VERSION : 0.1
   VAR_INPUT
      Nr_Ost_Elementu : Int;   // Numer ostatniego elementu, dla ktorego wykonywana jest klasa
      Nr_Plc : Byte;
   END_VAR
   VAR_TEMP
      i : Int;
   END_VAR
BEGIN
   FOR #i := 1 TO #Nr_Ost_Elementu BY 1 DO
       REGION Opisy bitow sygnalow: bRoz,bSym,bSt,bSt_1,bTrP
           //bRoz - ROZKAZ OPERATORA - DB322.DBW10 - WORD
           //bRozB1
           //"DB322_DV1".DV1[#i].bRoZB1.%X0 - Tryb pracy: 0-Zdalny reczny; 1-Zdalny auto
           //"DB322_DV1".DV1[#i].bRoZB1.%X1 - Symulacja wejsc urz: 0-Wylaczona; 1-Zalaczona
           //"DB322_DV1".DV1[#i].bRoZB1.%X2 - Praca z wyjsciami urz: 0-Wylaczona; 1-Zalaczona
           //"DB322_DV1".DV1[#i].bRoZB1.%X3 - Sterowanie urz. w tr. Zdalnym-Man: 0-Wylacz; 1-Zalacz
           //"DB322_DV1".DV1[#i].bRoZB1.%X4 - Sterowanie kier. w tr. Zdalnym-Man: 0-Lewa; 1-Prawo
           //"DB322_DV1".DV1[#i].bRoZB1.%X5 - Rezerwa
           //"DB322_DV1".DV1[#i].bRoZB1.%X6 - Monitoring potwierdzen zal/wyl: 0-Wylaczone; 1-Zalaczone
           //"DB322_DV1".DV1[#i].bRoZB1.%X7 - Rezerwa
           //bRozB2
           //"DB322_DV1".DV1[#i].bRoZB2.%X0 - Kasuj awarie (impuls)
           //"DB322_DV1".DV1[#i].bRoZB2.%X1-X7 - Rezerwa (impuls)
           //
           //bSym - SYM WEJSCIA - DB322.DBW12 - WORD
           //"DB322_DV1".DV1[#i].bSym.%X0 - Aktywacja urz. w systemie (ustawiany tylko z programu)
           //"DB322_DV1".DV1[#i].bSym.%X1 - Sterowanie urz. w tr. Zdalnym-Auto: 0-Wylacz; 1-Zalacz
           //"DB322_DV1".DV1[#i].bSym.%X2 - Potwierdzenie zalaczenia/otwarcia
           //"DB322_DV1".DV1[#i].bSym.%X3 - Potwierdzenie wylaczenia/zamkniecia
           //"DB322_DV1".DV1[#i].bSym.%X4 - Potwierdzenie gotowosci
           //"DB322_DV1".DV1[#i].bSym.%X5 - Tryb sterowania: 0-Zdalne z PC; 1-Lokalne z elewacji szafy
           //"DB322_DV1".DV1[#i].bSym.%X6 - Tryb remontowy (z wylacznika): 0-Brak; 1-Aktywny
           //"DB322_DV1".DV1[#i].bSym.%X7 - Awaria zewnetrzna: 0-Brak; 1-Aktywny
           //"DB322_DV1".DV1[#i].bSym.%X8 - Blokada zmiany tr. zdalnego z Auto na Man: 0-Brak; 1-Aktywna
           //"DB322_DV1".DV1[#i].bSym.%X9 - Interlock w trybie Zdalnym-Auto: 0-Brak; 1-Aktywny
           //"DB322_DV1".DV1[#i].bSym.%X10-X15 - Rezerwa
           //
           //bSt_Tryb - STAN - DB322.DBW14 - WORD
           //"DB322_DV1".DV1[#i].bSt_Tryb.%X0 - Awaria od braku potwierdzen: 0-Nieaktywna; 1-Aktywna
           //"DB322_DV1".DV1[#i].bSt_Tryb.%X1 - Awaria od braku gotowosci: 0-Nieaktywna; 1-Aktywna
           //"DB322_DV1".DV1[#i].bSt_Tryb.%X2 - Awaria zewnetzrna: 0-Nieaktywna; 1-Aktywna
           //"DB322_DV1".DV1[#i].bSt_Tryb.%X3-X6 - Awaria rezerwa
           //"DB322_DV1".DV1[#i].bSt_Tryb.%X7 - Monitoring potwierdzen: 0-Wylaczony; 1-Zalaczony
           //"DB322_DV1".DV1[#i].bSt_Tryb.%X8 - Urzadzenie aktywowane
           //"DB322_DV1".DV1[#i].bSt_Tryb.%X9 - Blokada zmaiany tr. zdalnego z Auto na Man: 0-Brak; 1-Aktywna
           //"DB322_DV1".DV1[#i].bSt_Tryb.%X10 - Stan wyjścia sterującego obiekt: 0-Zamknij; 1-Otwórz
           //"DB322_DV1".DV1[#i].bSt_Tryb.%X11 - Interlock w trybie Zdalnym-Auto: 0-Brak; 1-Aktywny
           //"DB322_DV1".DV1[#i].bSt_Tryb.%X12 - Symulacja wejsc urzadzenia: 0-Wylaczona; 1-Zalaczona
           //"DB322_DV1".DV1[#i].bSt_Tryb.%X13 - Praca z wyjsciami urzadzenia: 0-Wylaczona; 1-Zalaczona
           //"DB322_DV1".DV1[#i].bSt_Tryb.%X14 - Stan urzadzenia: 0-Brak odliczania czasu do otwarcia 1-Odliczanie
           //"DB322_DV1".DV1[#i].bSt_Tryb.%X15 - Stan urzadzenia: 0-Brak odliczania czasu do zamkniecia 1-Odliczanie
           //
           //bSt_Urz - STAN - DB322.DBW16 - INT
           //"DB322_DV1".DV1[#i].bSt_Urz.%X0 - STAN(1)- Awaria zbiorcza 1-Aktywna; 0-Brak aktywnosci obiektu
           //"DB322_DV1".DV1[#i].bSt_Urz.%X1 - STAN(2)- Urzadzenie: 1-Zamkniete; 0-Inny stan
           //"DB322_DV1".DV1[#i].bSt_Urz.%X2 - STAN(4)- Urzadzenie: 1-Otwieranie; 0-Inny stan
           //"DB322_DV1".DV1[#i].bSt_Urz.%X3 - STAN(8)- Urzadzenie: 1-Otwarte; 0-Inny stan
           //"DB322_DV1".DV1[#i].bSt_Urz.%X4 - STAN(16)- Urzadzenie: 1-Zamykanie; 0-Inny stan
           //"DB322_DV1".DV1[#i].bSt_Urz.%X5 - STAN(32)- Urzadzenie: 1-Odliczanie czasu zwloki awarii; 0-Inny stan
           //"DB322_DV1".DV1[#i].bSt_Urz.%X6-X7 - STAN- Stan rezerwa
           //
           //bTrP - TRYB PRACY - DB322.DBW17 - INT
           //"DB322_DV1".DV1[#i].bTrP.%X0 - TRYB PRACY(1) - Tryb Remontowy(1): 1-Aktywny; 0-Brak aktywnosci obiektu
           //"DB322_DV1".DV1[#i].bTrP.%X1 - Tryb PRACY(2) - Tryb Sterowania: 1-Lokalny - z szafy; 0-Inny stan
           //"DB322_DV1".DV1[#i].bTrP.%X2 - TRYB PRACY(4) - Tryb Sterowania Zdalnego: 1-Zdalny Reczny; 0-Inny stan
           //"DB322_DV1".DV1[#i].bTrP.%X3 - TRYB PRACY(8) - Tryb Sterowania Zdalnego: 1-Zdalny Automatyczny; 0-Inny stan
           //"DB322_DV1".DV1[#i].bTrP.%X4-X7 - Tryb PRACY(16)(32)(64)(128): Rezerwa
       END_REGION
       REGION Przepisanie danych do obiektu
           "DB322_DV1".DV1[#i].yNrID := #i;
           "DB322_DV1".DV1[#i].yNrPLC := #Nr_Plc;
       END_REGION
       REGION Warunek na wykonanie funkcji
           "DB322_DV1".DV1[#i].bSym.%X0 := "DB322_DV1".DV1[#i].bWeAkt;
           IF "DB322_DV1".DV1[#i].bWeAkt = 0 THEN //Akcja przy deaktywowaniu obiektu
               "DB322_DV1".DV1[#i].bWeZalAuto := 0;
               "DB322_DV1".DV1[#i].bWePotwZal := 0;
               "DB322_DV1".DV1[#i].bWePotwWyl := 0;
               "DB322_DV1".DV1[#i].bWePotwGot := 0;
               "DB322_DV1".DV1[#i].bWeTrRem := 0;
               "DB322_DV1".DV1[#i].bWeAwrZ := 0;
               "DB322_DV1".DV1[#i].bWeBlZmAuto := 0;
               "DB322_DV1".DV1[#i].bWeIlock := 0;
               "DB322_DV1".DV1[#i].bRoZB1 := 0;
               "DB322_DV1".DV1[#i].bRoZB2 := 0;
               "DB322_DV1".DV1[#i].bSym := 0;
               "DB322_DV1".DV1[#i].bSt_Tryb := 0;
               "DB322_DV1".DV1[#i].bSt_Urz := 0;
               "DB322_DV1".DV1[#i].bTrP := 0;
               "DB322_DV1".DV1[#i].bWySter := 0;
               "DB322_DV1".DV1[#i].bWyRst := 0;
           ELSE
               REGION Program funckji
                   REGION Symulacja wejsc - przepisywanie wartosci wejsciowych, gdy nie ma symulacji oprocz bWeAkt
                       IF "DB322_DV1".DV1[#i].bSt_Tryb.%X12 = 0 THEN
                           "DB322_DV1".DV1[#i].bSym.%X1 := "DB322_DV1".DV1[#i].bWeZalAuto;
                           "DB322_DV1".DV1[#i].bSym.%X2 := "DB322_DV1".DV1[#i].bWePotwZal;
                           "DB322_DV1".DV1[#i].bSym.%X3 := "DB322_DV1".DV1[#i].bWePotwWyl;
                           "DB322_DV1".DV1[#i].bSym.%X4 := "DB322_DV1".DV1[#i].bWePotwGot;
                           "DB322_DV1".DV1[#i].bSym.%X5 := "DB322_DV1".DV1[#i].bWeTrLok;
                           "DB322_DV1".DV1[#i].bSym.%X6 := "DB322_DV1".DV1[#i].bWeTrRem;
                           "DB322_DV1".DV1[#i].bSym.%X7 := "DB322_DV1".DV1[#i].bWeAwrZ;
                           "DB322_DV1".DV1[#i].bSym.%X8 := "DB322_DV1".DV1[#i].bWeBlZmAuto;
                           "DB322_DV1".DV1[#i].bSym.%X9 := "DB322_DV1".DV1[#i].bWeIlock;
                       END_IF;
                   END_REGION
                   REGION Okreslenie stanow    
                       "DB322_DV1".DV1[#i].bSt_Tryb.%X7 := "DB322_DV1".DV1[#i].bRoZB1.%X6;
                       "DB322_DV1".DV1[#i].bSt_Tryb.%X8 := "DB322_DV1".DV1[#i].bWeAkt;
                       "DB322_DV1".DV1[#i].bSt_Tryb.%X9 := (("DB322_DV1".DV1[#i].bSym.%X8 AND "DB322_DV1".DV1[#i].bSt_Tryb.%X12) OR ("DB322_DV1".DV1[#i].bWeBlZmAuto AND NOT "DB322_DV1".DV1[#i].bSt_Tryb.%X12));
                       "DB322_DV1".DV1[#i].bSt_Tryb.%X10 := "DB322_DV1".DV1[#i].bHlp186 AND "DB322_DV1".DV1[#i].bSt_Tryb.%X13;
                       "DB322_DV1".DV1[#i].bSt_Tryb.%X11 := (("DB322_DV1".DV1[#i].bSym.%X9 AND "DB322_DV1".DV1[#i].bSt_Tryb.%X12) OR ("DB322_DV1".DV1[#i].bWeIlock AND NOT "DB322_DV1".DV1[#i].bSt_Tryb.%X12));
                       "DB322_DV1".DV1[#i].bSt_Tryb.%X12 := "DB322_DV1".DV1[#i].bRoZB1.%X1;
                       "DB322_DV1".DV1[#i].bSt_Tryb.%X13 := "DB322_DV1".DV1[#i].bRoZB1.%X2;
                   END_REGION
                   REGION Filtracja
                       REGION Timer 1,2 - opoznienie zalaczenia i wylaczenia
                           "DB322_DV1".DV1[#i].bTmr_On_Start := ("DB322_DV1".DV1[#i].bSym.%X1 AND "DB322_DV1".DV1[#i].bSt_Tryb.%X12) OR ("DB322_DV1".DV1[#i].bWeZalAuto AND NOT "DB322_DV1".DV1[#i].bSt_Tryb.%X12);
                           "DB322_DV1".DV1[#i].bTmr_Off_Start := NOT (("DB322_DV1".DV1[#i].bSym.%X1 AND "DB322_DV1".DV1[#i].bSt_Tryb.%X12) OR ("DB322_DV1".DV1[#i].bWeZalAuto AND NOT "DB322_DV1".DV1[#i].bSt_Tryb.%X12));
                           "FC301_Timer"(iTyp := 1,
                                         bOnOff := "DB322_DV1".DV1[#i].bTmr_On_Start,
                                         bRst := 0,
                                         dCzasZad := "DB322_DV1".DV1[#i].yCzZadOpzZal,
                                         timer_1s := "imp1s",
                                         bOk => "DB322_DV1".DV1[#i].bTmr_On_Ok,
                                         dCzasAkt := "DB322_DV1".DV1[#i].yCzAktOpzZal);
                           "FC301_Timer"(iTyp := 1,
                                         bOnOff := "DB322_DV1".DV1[#i].bTmr_Off_Start,
                                         bRst := 0,
                                         dCzasZad := "DB322_DV1".DV1[#i].yCzZadOpzWyl,
                                         timer_1s := "imp1s",
                                         bOk => "DB322_DV1".DV1[#i].bTmr_Off_Ok,
                                         dCzasAkt := "DB322_DV1".DV1[#i].yCzAktOpzWyl);

                       END_REGION
                       REGION Efekt dzialania timerow - blok NoNc
                           // zmiana aby nie zamykal zaworu przy awarii
                           IF "DB322_DV1".DV1[#i].bTmr_On_Ok THEN
                               "DB322_DV1".DV1[#i].bHlp184 := 1;
                           END_IF;
                           IF "DB322_DV1".DV1[#i].bTmr_Off_Ok THEN //OR "DB322_DV1".DV1[#i].bSt_Urz = 1 THEN
                               "DB322_DV1".DV1[#i].bHlp184 := 0;
                           END_IF;

                           IF "DB322_DV1".DV1[#i].bTmr_Off_Ok THEN
                               "DB322_DV1".DV1[#i].bHlp185 := 1;
                           END_IF;
                           IF "DB322_DV1".DV1[#i].bTmr_On_Ok THEN //OR "DB322_DV1".DV1[#i].bSt_Urz = 1 THEN
                               "DB322_DV1".DV1[#i].bHlp185 := 0;
                           END_IF;

                           "DB322_DV1".DV1[#i].bHlp187 := (NOT "DB322_DV1".DV1[#i].bNoNc AND "DB322_DV1".DV1[#i].bHlp184) OR ("DB322_DV1".DV1[#i].bNoNc AND "DB322_DV1".DV1[#i].bHlp185);
                       END_REGION
                       REGION Stany zaworu przy odliczaniu czasu
                           "DB322_DV1".DV1[#i].bSt_Tryb.%X14 := "DB322_DV1".DV1[#i].bTmr_On_Start AND NOT "DB322_DV1".DV1[#i].bTmr_On_Ok;
                           "DB322_DV1".DV1[#i].bSt_Tryb.%X15 := ("DB322_DV1".DV1[#i].bTmr_Off_Start AND NOT "DB322_DV1".DV1[#i].bTmr_Off_Ok);
                       END_REGION
                   END_REGION
                   REGION Generowanie sygnalu alarmu 
                       REGION Zerowanie czasu awarii przy zmianie sterowania podczas ruchu
                           "R_TRIG_DB_6"(CLK := "DB322_DV1".DV1[#i].bHlp186 AND "DB322_DV1".DV1[#i].bSt_Urz <> 1,
                                         Q => "DB322_DV1".DV1[#i].bHlp256);
                           "R_TRIG_DB"(CLK:=NOT "DB322_DV1".DV1[#i].bHlp186 AND "DB322_DV1".DV1[#i].bSt_Urz <> 1,
                                       Q=>"DB322_DV1".DV1[#i].bHlp257);

                           IF "DB322_DV1".DV1[#i].bHlp256 OR "DB322_DV1".DV1[#i].bHlp257 THEN
                               "DB322_DV1".DV1[#i].yCzasAktOpzAlm := 0;
                           END_IF;
                       END_REGION
                       REGION Sygnal bledu od potwierdzen.
                           // Jezeli brak bitu monitoringu lub bitu pracy z wyjsciami nie ma awarii. Jezeli jest tryb lokalny lub remontowy nie ma awarii
                           "DB322_DV1".DV1[#i].bHlp_NoNc := "DB322_DV1".DV1[#i].bNoNc XOR "DB322_DV1".DV1[#i].bHlp186;

                           "DB322_DV1".DV1[#i].bTmr_Awr_Start := (("DB322_DV1".DV1[#i].bHlp_NoNc XOR (("DB322_DV1".DV1[#i].bWePotwZal AND NOT "DB322_DV1".DV1[#i].bSt_Tryb.%X12) OR ("DB322_DV1".DV1[#i].bSym.%X2 AND "DB322_DV1".DV1[#i].bSt_Tryb.%X12))))
                           OR (NOT "DB322_DV1".DV1[#i].bHlp_NoNc AND NOT (("DB322_DV1".DV1[#i].bWePotwWyl AND NOT "DB322_DV1".DV1[#i].bSt_Tryb.%X12) OR ("DB322_DV1".DV1[#i].bSym.%X3 AND "DB322_DV1".DV1[#i].bSt_Tryb.%X12)))
                           OR ("DB322_DV1".DV1[#i].bHlp_NoNc AND ("DB322_DV1".DV1[#i].bWePotwWyl AND NOT "DB322_DV1".DV1[#i].bSt_Tryb.%X12) OR ("DB322_DV1".DV1[#i].bSym.%X3 AND "DB322_DV1".DV1[#i].bSt_Tryb.%X12))
                           OR ((("DB322_DV1".DV1[#i].bWePotwZal AND NOT "DB322_DV1".DV1[#i].bSt_Tryb.%X12) OR ("DB322_DV1".DV1[#i].bSym.%X2 AND "DB322_DV1".DV1[#i].bSt_Tryb.%X12)) AND (("DB322_DV1".DV1[#i].bWePotwWyl AND NOT "DB322_DV1".DV1[#i].bSt_Tryb.%X12) OR ("DB322_DV1".DV1[#i].bSym.%X3 AND "DB322_DV1".DV1[#i].bSt_Tryb.%X12)))
                           OR (NOT (("DB322_DV1".DV1[#i].bWePotwZal AND NOT "DB322_DV1".DV1[#i].bSt_Tryb.%X12) OR ("DB322_DV1".DV1[#i].bSym.%X2 AND "DB322_DV1".DV1[#i].bSt_Tryb.%X12)) AND (NOT ("DB322_DV1".DV1[#i].bWePotwWyl AND NOT "DB322_DV1".DV1[#i].bSt_Tryb.%X12) OR ("DB322_DV1".DV1[#i].bSym.%X3 AND "DB322_DV1".DV1[#i].bSt_Tryb.%X12)))
                           AND "DB322_DV1".DV1[#i].bSt_Tryb.%X7 AND "DB322_DV1".DV1[#i].bSt_Tryb.%X13 AND "DB322_DV1".DV1[#i].bTrP <> 1 AND "DB322_DV1".DV1[#i].bTrP <> 2 AND NOT "DB322_DV1".DV1[#i].bRoZB2.%X0;

                       END_REGION
                       REGION Timer 3 - kontrola alarmu
                           "FC301_Timer"(iTyp := 1,
                                         bOnOff := "DB322_DV1".DV1[#i].bTmr_Awr_Start,
                                         bRst := 0,
                                         dCzasZad := "DB322_DV1".DV1[#i].yCzZadOpzAlm,
                                         timer_1s := "imp1s",
                                         bOk => "DB322_DV1".DV1[#i].bTmr_Alm_Ok,
                                         dCzasAkt := "DB322_DV1".DV1[#i].yCzasAktOpzAlm);


                       END_REGION
                       REGION Ustawienie i kasowanie sygnalu awarii
                           IF "DB322_DV1".DV1[#i].bTmr_Alm_Ok THEN
                               "DB322_DV1".DV1[#i].bSt_Tryb.%X0 := 1
                               ;
                           END_IF;
                           IF NOT (("DB322_DV1".DV1[#i].bWePotwGot AND NOT "DB322_DV1".DV1[#i].bSt_Tryb.%X12) OR ("DB322_DV1".DV1[#i].bSym.%X4 AND "DB322_DV1".DV1[#i].bSt_Tryb.%X12)) THEN
                               "DB322_DV1".DV1[#i].bSt_Tryb.%X1 := 1
                               ;
                           END_IF;
                           IF ("DB322_DV1".DV1[#i].bWeAwrZ AND NOT "DB322_DV1".DV1[#i].bSt_Tryb.%X12) OR ("DB322_DV1".DV1[#i].bSym.%X7 AND "DB322_DV1".DV1[#i].bSt_Tryb.%X12) THEN
                               "DB322_DV1".DV1[#i].bSt_Tryb.%X2 := 1
                               ;
                           END_IF;
                           IF "DB322_DV1".DV1[#i].bRoZB2.%X0 AND "DB322_DV1".DV1[#i].bSt_Urz=1 THEN //zmiana 2.10.23 - reset tylko obiektu w awarii
                               "DB322_DV1".DV1[#i].bSt_Tryb := 0
                               ;
                           END_IF;
                       END_REGION
                   END_REGION
                   REGION Tryb pracy i sterowanie wyjsciem
                       REGION Przepisanie potwierdzen na sterowanie reczne gdy tryb lokalny
                           // Przypadek gdy ktos z wlaczonym lokalnie urz. przechodzi na tryb zdalny-reczny
                           IF "DB322_DV1".DV1[#i].bTrP = 2 THEN

                               "DB322_DV1".DV1[#i].bRoZB1.%X0 := 0;

                               IF (("DB322_DV1".DV1[#i].bWePotwWyl AND NOT "DB322_DV1".DV1[#i].bSt_Tryb.%X12) OR ("DB322_DV1".DV1[#i].bSym.%X3 AND "DB322_DV1".DV1[#i].bSt_Tryb.%X12)) THEN
                                   "DB322_DV1".DV1[#i].bRoZB1.%X3 := 0;
                               END_IF;

                               IF (("DB322_DV1".DV1[#i].bWePotwZal AND NOT "DB322_DV1".DV1[#i].bSt_Tryb.%X12) OR ("DB322_DV1".DV1[#i].bSym.%X2 AND "DB322_DV1".DV1[#i].bSt_Tryb.%X12)) THEN
                                   "DB322_DV1".DV1[#i].bRoZB1.%X3 := 1
                                   ;
                               END_IF;
                               ;
                           END_IF;

                       END_REGION
                       REGION Przepisanie potwierdzen na sterowanie reczne gdy tryb zdalny-auto
                           // Przypadek gdy ktos z wlaczonym automatycznie urz. przechodzi na tryb zdalny-reczny
                           IF "DB322_DV1".DV1[#i].bTrP = 8 THEN
                               "DB322_DV1".DV1[#i].bRoZB1.%X3 :=(("DB322_DV1".DV1[#i].bWeZalAuto AND NOT "DB322_DV1".DV1[#i].bSt_Tryb.%X12) OR ("DB322_DV1".DV1[#i].bSym.%X1 AND "DB322_DV1".DV1[#i].bSt_Tryb.%X12));
                               ;
                           END_IF;


                       END_REGION
                       REGION Blokada zmiany trybu zdalny-automatyczny
                           IF "DB322_DV1".DV1[#i].bTrP = 8 AND "DB322_DV1".DV1[#i].bSt_Tryb.%X9 THEN
                               "DB322_DV1".DV1[#i].bRoZB1.%X0 := 1;
                               ;
                           END_IF;
                       END_REGION
                       REGION Blokada zalaczenia urzadzenia w trybie zdalnym-manualnym przy zalaczonym Interlocku
                           IF "DB322_DV1".DV1[#i].bWeIlock THEN
                               "DB322_DV1".DV1[#i].bRoZB1.%X3 := 0;
                           END_IF;

                       END_REGION
                       REGION Okreslenie trybu pracy wyjscia
                           IF  "DB322_DV1".DV1[#i].bRoZB1.%X0 AND NOT "DB322_DV1".DV1[#i].bSt_Tryb.%X9 THEN
                               "DB322_DV1".DV1[#i].bTrP := 8
                               ;
                           END_IF;
                           IF NOT "DB322_DV1".DV1[#i].bRoZB1.%X0 THEN
                               "DB322_DV1".DV1[#i].bTrP := 4
                               ;
                           END_IF;
                           IF ("DB322_DV1".DV1[#i].bWeTrLok AND NOT "DB322_DV1".DV1[#i].bSt_Tryb.%X12) OR ("DB322_DV1".DV1[#i].bSym.%X5 AND "DB322_DV1".DV1[#i].bSt_Tryb.%X12) THEN
                               "DB322_DV1".DV1[#i].bTrP := 2
                               ;
                           END_IF;
                           IF ("DB322_DV1".DV1[#i].bWeTrRem AND NOT "DB322_DV1".DV1[#i].bSt_Tryb.%X12) OR ("DB322_DV1".DV1[#i].bSym.%X6 AND "DB322_DV1".DV1[#i].bSt_Tryb.%X12) THEN
                               "DB322_DV1".DV1[#i].bTrP := 1
                               ;
                           END_IF;
                       END_REGION
                       REGION Sterowanie wyjsciem
                           // zmiana - ignorowanie awarii - brak zmiany stanu wyjscia
                           "DB322_DV1".DV1[#i].bHlp186 := (("DB322_DV1".DV1[#i].bTrP = 8 AND "DB322_DV1".DV1[#i].bHlp187) OR ("DB322_DV1".DV1[#i].bTrP = 4 AND ("DB322_DV1".DV1[#i].bRoZB1.%X3 XOR "DB322_DV1".DV1[#i].bNoNc)))
                           AND NOT (("DB322_DV1".DV1[#i].bWeIlock AND NOT "DB322_DV1".DV1[#i].bSt_Tryb.%X12) OR ("DB322_DV1".DV1[#i].bSym.%X9 AND "DB322_DV1".DV1[#i].bSt_Tryb.%X12));// AND "DB322_DV1".DV1[#i].bSt_Urz <> 1;
                           "DB322_DV1".DV1[#i].bWySter:= "DB322_DV1".DV1[#i].bHlp186 AND "DB322_DV1".DV1[#i].bSt_Tryb.%X13;
                       END_REGION
                       REGION Sterowanie resetem
                           "DB322_DV1".DV1[#i].bWyRst := "DB322_DV1".DV1[#i].bRoZB2.%X0;
                        END_REGION
                       REGION Stan urzadzenia
                           "DB322_DV1".DV1[#i].bSt_Urz := 0; //czyszczenie stanu
                           REGION Urzadzenie otwierane
                               //kazda inna kombinacja potwierdzen niz przy urz. "otwartym"
                               IF "DB322_DV1".DV1[#i].bSt_Tryb.%X7 AND "DB322_DV1".DV1[#i].bSt_Tryb.%X13 AND "DB322_DV1".DV1[#i].bHlp_NoNc THEN
                                   "DB322_DV1".DV1[#i].bSt_Urz := 4
                                   ;
                               END_IF;

                           END_REGION
                           REGION Urzadzenie zamykane
                               // kazda inna kombinacja potwierdzen niz przy urz. zamknietym
                               IF "DB322_DV1".DV1[#i].bSt_Tryb.%X7 AND "DB322_DV1".DV1[#i].bSt_Tryb.%X13 AND NOT "DB322_DV1".DV1[#i].bHlp_NoNc THEN
                                   "DB322_DV1".DV1[#i].bSt_Urz := 16
                                   ;
                               END_IF;
                           END_REGION
                           REGION Urzadzenie zamkniete
                               IF "DB322_DV1".DV1[#i].bTrP <> 2 AND (("DB322_DV1".DV1[#i].bSt_Tryb.%X7 AND "DB322_DV1".DV1[#i].bSt_Tryb.%X13 AND NOT "DB322_DV1".DV1[#i].bHlp_NoNc
                                   AND (("DB322_DV1".DV1[#i].bWePotwWyl AND NOT "DB322_DV1".DV1[#i].bSt_Tryb.%X12) OR ("DB322_DV1".DV1[#i].bSym.%X3 AND "DB322_DV1".DV1[#i].bSt_Tryb.%X12))
                                   AND NOT (("DB322_DV1".DV1[#i].bWePotwZal AND NOT "DB322_DV1".DV1[#i].bSt_Tryb.%X12) OR ("DB322_DV1".DV1[#i].bSym.%X2 AND "DB322_DV1".DV1[#i].bSt_Tryb.%X12)))
                                   OR (NOT "DB322_DV1".DV1[#i].bSt_Tryb.%X7 OR NOT "DB322_DV1".DV1[#i].bSt_Tryb.%X13) AND NOT "DB322_DV1".DV1[#i].bHlp186)
                                   OR (("DB322_DV1".DV1[#i].bTrP = 2 AND (("DB322_DV1".DV1[#i].bWePotwWyl AND NOT "DB322_DV1".DV1[#i].bSt_Tryb.%X12) OR ("DB322_DV1".DV1[#i].bSym.%X3 AND "DB322_DV1".DV1[#i].bSt_Tryb.%X12))) OR "DB322_DV1".DV1[#i].bTrP = 1)
                               THEN
                                   "DB322_DV1".DV1[#i].bSt_Urz := 2 //Urzadzenie zamkniete
                                   ;
                               END_IF;
                           END_REGION
                           REGION Urzadzenie otwarte
                               IF "DB322_DV1".DV1[#i].bTrP <> 2 AND (("DB322_DV1".DV1[#i].bSt_Tryb.%X7 AND "DB322_DV1".DV1[#i].bSt_Tryb.%X13 AND "DB322_DV1".DV1[#i].bHlp_NoNc
                                   AND NOT (("DB322_DV1".DV1[#i].bWePotwWyl AND NOT "DB322_DV1".DV1[#i].bSt_Tryb.%X12) OR ("DB322_DV1".DV1[#i].bSym.%X3 AND "DB322_DV1".DV1[#i].bSt_Tryb.%X12))
                                   AND (("DB322_DV1".DV1[#i].bWePotwZal AND NOT "DB322_DV1".DV1[#i].bSt_Tryb.%X12) OR ("DB322_DV1".DV1[#i].bSym.%X2 AND "DB322_DV1".DV1[#i].bSt_Tryb.%X12)))
                                   OR (NOT "DB322_DV1".DV1[#i].bSt_Tryb.%X7 OR NOT "DB322_DV1".DV1[#i].bSt_Tryb.%X13) AND "DB322_DV1".DV1[#i].bHlp186)
                                   OR ("DB322_DV1".DV1[#i].bTrP = 2 AND ("DB322_DV1".DV1[#i].bWePotwZal OR "DB322_DV1".DV1[#i].bSym.%X2))
                               THEN
                                   "DB322_DV1".DV1[#i].bSt_Urz := 8  //Urzadzenie otwarte
                                   ;
                               END_IF;
                           END_REGION
                           REGION Awaria zbiorcza
                               IF "DB322_DV1".DV1[#i].bSt_Tryb.%X0 OR "DB322_DV1".DV1[#i].bSt_Tryb.%X1 OR "DB322_DV1".DV1[#i].bSt_Tryb.%X2 THEN
                                   "DB322_DV1".DV1[#i].bSt_Urz := 1 //Awaria zbiorcza
                                   ;
                               END_IF;
                           END_REGION



                       END_REGION
                   END_REGION
                   REGION Ustawienia koncowe
                       // Samokasowanie sygnalow
                       "DB322_DV1".DV1[#i].bRoZB2 := 0;
                       IF "DB322_DV1".DV1[#i].bAoff = 1 THEN
                           "DB322_DV1".DV1[#i].bWeZalAuto := 0;
                       END_IF;
                   END_REGION
               END_REGION
           END_IF;
       END_REGION
   END_FOR;
END_FUNCTION

FUNCTION "FC323_DM1" : Void   // FC323, SCL
{ S7_Optimized_Access := 'TRUE' }
VERSION : 0.1
   VAR_INPUT
      Nr_Ost_Elementu : Int;   // Numer ostatniego elementu, dla ktorego wykonywana jest klasa
      Nr_Plc : Byte;
      bKier : Bool;   // Bit wyboru stacyjki: 0-Bez kierunku; 1-Z kierunkiem
   END_VAR
   VAR_TEMP
      i : Int;
   END_VAR
BEGIN
   FOR #i := 1 TO #Nr_Ost_Elementu BY 1 DO
       REGION Opisy bitow sygnalow: bRoz,bSym,bSt,bSt_1,bTrP
           //bRoz - ROZKAZ OPERATORA - DB323.DBW10 - WORD
           //bRozB1
           //"DB323_DM1".DM1[#i].bRoZB1.%X0 - Tryb pracy: 0-Zdalny reczny; 1-Zdalny auto
           //"DB323_DM1".DM1[#i].bRoZB1.%X1 - Symulacja wejsc urz: 0-Wylaczona; 1-Zalaczona
           //"DB323_DM1".DM1[#i].bRoZB1.%X2 - Praca z wyjsciami urz: 0-Wylaczona; 1-Zalaczona
           //"DB323_DM1".DM1[#i].bRoZB1.%X3 - Sterowanie urz. w tr. Zdalnym-Man: 0-Wylacz; 1-Zalacz
           //"DB323_DM1".DM1[#i].bRoZB1.%X4 - Sterowanie kier. w tr. Zdalnym-Man: 0-Lewa; 1-Prawo
           //"DB323_DM1".DM1[#i].bRoZB1.%X5 - Rezerwa
           //"DB323_DM1".DM1[#i].bRoZB1.%X6 - Monitoring potwierdzen zal/wyl: 0-Wylaczone; 1-Zalaczone
           //"DB323_DM1".DM1[#i].bRoZB1.%X7 - Rezerwa
           //bRozB2
           //"DB323_DM1".DM1[#i].bRoZB2.%X0 - Kasuj awarie (impuls)
           //"DB323_DM1".DM1[#i].bRoZB2.%X1-X7 - Rezerwa (impuls)
           //
           //bSym - SYM WEJSCIA - DB323.DBW12 - WORD
           //"DB323_DM1".DM1[#i].bSym.%X0 - Aktywacja urz. w systemie (ustawiany tylko z programu)
           //"DB323_DM1".DM1[#i].bSym.%X1 - Sterowanie urz. w tr. Zdalnym-Auto: 0-Wylacz; 1-Zalacz
           //"DB323_DM1".DM1[#i].bSym.%X2 - Potwierdzenie zalaczenia/otwarcia
           //"DB323_DM1".DM1[#i].bSym.%X3 - Potwierdzenie wylaczenia/zamkniecia
           //"DB323_DM1".DM1[#i].bSym.%X4 - Potwierdzenie gotowosci
           //"DB323_DM1".DM1[#i].bSym.%X5 - Tryb sterowania: 0-Zdalne z PC; 1-Lokalne z elewacji szafy
           //"DB323_DM1".DM1[#i].bSym.%X6 - Tryb remontowy (z wylacznika): 0-Brak; 1-Aktywny
           //"DB323_DM1".DM1[#i].bSym.%X7 - Awaria zewnetrzna: 0-Brak; 1-Aktywny
           //"DB323_DM1".DM1[#i].bSym.%X8 - Blokada zmiany tr. zdalnego z Auto na Man: 0-Brak; 1-Aktywna
           //"DB323_DM1".DM1[#i].bSym.%X9 - Interlock w trybie Zdalnym-Auto: 0-Brak; 1-Aktywny
           //"DB323_DM1".DM1[#i].bSym.%X10 - Kierunek obrotow: 0-Prawo; 1-Lewo
           //"DB323_DM1".DM1[#i].bSym.%X11-X15 - Rezerwa
           //
           //bSt_Tryb - STAN - DB323.DBW14 - WORD
           //"DB323_DM1".DM1[#i].bSt_Tryb.%X0 - Awaria od braku potwierdzen: 0-Nieaktywna; 1-Aktywna
           //"DB323_DM1".DM1[#i].bSt_Tryb.%X1 - Awaria od braku gotowosci: 0-Nieaktywna; 1-Aktywna
           //"DB323_DM1".DM1[#i].bSt_Tryb.%X2 - Awaria zewnetzrna: 0-Nieaktywna; 1-Aktywna
           //"DB323_DM1".DM1[#i].bSt_Tryb.%X3-X6 - Awaria rezerwa
           //"DB323_DM1".DM1[#i].bSt_Tryb.%X7 - Monitoring potwierdzen: 0-Wylaczony; 1-Zalaczony
           //"DB323_DM1".DM1[#i].bSt_Tryb.%X8 - Urzadzenie aktywowane
           //"DB323_DM1".DM1[#i].bSt_Tryb.%X9 - Blokada zmaiany tr. zdalnego z Auto na Man: 0-Brak; 1-Aktywna
           //"DB323_DM1".DM1[#i].bSt_Tryb.%X10 - Kierunek urzadzenia: 0-Prawo; 1-Lewo
           //"DB323_DM1".DM1[#i].bSt_Tryb.%X11 - Interlock w trybie Zdalnym-Auto: 0-Brak; 1-Aktywny